screen "Dev_AI" 800x480, template "Settings"
   Softkey "Softkey_F3" at 0,0 size 0x0
      on KeyDown: function_dd21b452("AI_x_Result", 1)
   Softkey "Softkey_F7" at 0,0 size 0x0
      on KeyDown: SetBit("AI_x_CMD_Reset")
   Button "Button_2" at 165,265 size 112x32; TextOff 'DB 300'; Authorization "User administration"
      on Release: SetTag("AIx", 300); SetTag("AIx_Name", 'DB 300')
      Visibility <- "Support_DB_All_AIs"
      Appearance <- "AIx"
   Button "Button_8" at 165,305 size 112x32; TextOff 'DB 301'; Authorization "User administration"
      on Release: SetTag("AIx", 301); SetTag("AIx_Name", 'DB 301')
      Visibility <- "Support_DB_All_AIs"
      Appearance <- "AIx"
   Button "Button_17" at 165,345 size 112x32; TextOff 'DB 302'; Authorization "User administration"
      on Release: SetTag("AIx", 302); SetTag("AIx_Name", 'DB 302')
      Visibility <- "Support_DB_All_AIs"
      Appearance <- "AIx"
   Button "Button_18" at 165,385 size 112x32; TextOff 'DB 303'; Authorization "User administration"
      on Release: SetTag("AIx", 303); SetTag("AIx_Name", 'DB 303')
      Visibility <- "Support_DB_All_AIs"
      Appearance <- "AIx"
   Button "Button_3" at 443,265 size 112x32; TextOff 'DB 310'; Authorization "User administration"
      on Release: SetTag("AIx", 310); SetTag("AIx_Name", 'DB 310')
      Visibility <- "Support_DB_All_AIs"
      Appearance <- "AIx"
   Button "Button_4" at 443,305 size 112x32; TextOff 'DB 311'; Authorization "User administration"
      on Release: SetTag("AIx", 311); SetTag("AIx_Name", 'DB 311')
      Visibility <- "Support_DB_All_AIs"
      Appearance <- "AIx"
   Button "Button_6" at 443,345 size 112x32; TextOff 'DB 312'; Authorization "User administration"
      on Release: SetTag("AIx", 312); SetTag("AIx_Name", 'DB 312')
      Visibility <- "Support_DB_All_AIs"
      Appearance <- "AIx"
   Button "Button_10" at 443,385 size 112x32; TextOff 'DB 313'; Authorization "User administration"
      on Release: SetTag("AIx", 313); SetTag("AIx_Name", 'DB 313')
      Visibility <- "Support_DB_All_AIs"
      Appearance <- "AIx"
   Button "Button_11" at 443,425 size 112x32; TextOff 'DB 314'; Authorization "User administration"
      on Release: SetTag("AIx", 314); SetTag("AIx_Name", 'DB 314')
      Visibility <- "Support_DB_All_AIs"
      Appearance <- "AIx"
   Button "Button_1" at 583,344 size 112x32; TextOff 'DB 317'; Authorization "User administration"
      on Release: SetTag("AIx", 317); SetTag("AIx_Name", 'DB 317')
      Visibility <- "Support_DB_All_AIs"
      Appearance <- "AIx"
   Button "Button_5" at 583,384 size 112x32; TextOff 'DB 318'; Authorization "User administration"
      on Release: SetTag("AIx", 318); SetTag("AIx_Name", 'DB 318')
      Visibility <- "Support_DB_All_AIs"
      Appearance <- "AIx"
   Button "Button_9" at 583,264 size 112x32; TextOff 'DB 315'; Authorization "User administration"
      on Release: SetTag("AIx", 315); SetTag("AIx_Name", 'DB 315')
      Visibility <- "Support_DB_All_AIs"
      Appearance <- "AIx"
   Button "Button_14" at 583,304 size 112x32; TextOff 'DB 316'; Authorization "User administration"
      on Release: SetTag("AIx", 316); SetTag("AIx_Name", 'DB 316')
      Visibility <- "Support_DB_All_AIs"
      Appearance <- "AIx"
   Rectangle "Rectangle_3" at 165,7 size 530x150
      Appearance <- "AI_x_CMD_Start_A"
   Button "Button_7" at 171,43 size 80x22; TextOff 'Авто'; Authorization "User administration"; TextList "Hand"
      on Click: InvertBit("AI_x_CMD_Hand")
      Appearance <- "AI_x_CMD_Hand"
      ProcessValue <- "AI_x_CMD_Hand"
   TextField "Text field_1" at 484,12 size 107x18; Text 'Масштабирование'
      Visibility <- "AI_x_Use_RTD"
   TextField "Text field_20" at 495,24 size 18x18; Text 'от'
      Visibility <- "AI_x_Use_RTD"
   IOField "I/O field_5" at 476,42 size 65x20; Authorization "User administration"; FormatPattern 99999
      ProcessValue <- "AI_x_Converter_Min_In"
      Visibility <- "AI_x_Use_RTD"
   TextField "Text field_21" at 559,24 size 19x18; Text 'до'
      Visibility <- "AI_x_Use_RTD"
   IOField "I/O field_11" at 171,82 size 80x30; Authorization "User administration"; FormatPattern s9999.9
      ProcessValue <- "AI_x_Result"
      Appearance <- "AI_x_Status"
   TextField "Text field_22" at 177,64 size 68x18; Text 'Показания:'
   TextField "Text field_23" at 180,113 size 63x18; Text 'Вход ПЛК:'
   IOField "I/O field_17" at 171,133 size 80x20; FormatPattern s99999
      ProcessValue <- "AI_x_Signal"
   TextField "Text field_24" at 489,89 size 42x18; Text 'Обрыв'
      Visibility <- "AI_x_Alarm_NC"
   TextField "Text field_25" at 555,89 size 42x18; Text 'КЗ'
      Visibility <- "AI_x_Alarm_SC"
   IOField "I/O field_18" at 544,42 size 65x20; Authorization "User administration"; FormatPattern 99999
      ProcessValue <- "AI_x_Converter_Max_In"
      Visibility <- "AI_x_Use_RTD"
   IOField "I/O field_24" at 476,66 size 65x20; Authorization "User administration"; FormatPattern s9999.99
      ProcessValue <- "AI_x_Converter_Min_Out"
      Visibility <- "AI_x_Use_RTD"
   IOField "I/O field_25" at 544,66 size 65x20; Authorization "User administration"; FormatPattern s9999.99
      ProcessValue <- "AI_x_Converter_Max_Out"
      Visibility <- "AI_x_Use_RTD"
   IOField "I/O field_10" at 382,35 size 55x20; Authorization "User administration"; FormatPattern s9999.9
      Appearance <- "AI_x_Alarm_HH"
      ProcessValue <- "AI_x_SP_HH"
   TextField "Text field_10" at 354,36 size 28x18; Text 'HHS'
   TextField "Text field_12" at 354,60 size 20x18; Text 'HS'
   IOField "I/O field_12" at 382,58 size 55x20; Authorization "User administration"; FormatPattern s9999.9
      Appearance <- "AI_x_Alarm_H"
      ProcessValue <- "AI_x_SP_H"
   IOField "I/O field_26" at 440,35 size 26x20; Authorization "User administration"; FormatPattern 99.9
      Appearance <- "AI_x_Alarm_HH"
      ProcessValue <- "AI_x_Timers_HH_SP"
   IOField "I/O field_27" at 440,58 size 26x20; Authorization "User administration"; FormatPattern 99.9
      Appearance <- "AI_x_Alarm_H"
      ProcessValue <- "AI_x_Timers_H_SP"
   IOField "I/O field_28" at 382,82 size 55x20; Authorization "User administration"; FormatPattern s9999.9
      Appearance <- "AI_x_Alarm_L"
      ProcessValue <- "AI_x_SP_L"
   TextField "Text field_6" at 354,84 size 18x18; Text 'LS'
   TextField "Text field_28" at 354,108 size 24x18; Text 'LLS'
   IOField "I/O field_29" at 382,106 size 55x20; Authorization "User administration"; FormatPattern s9999.9
      Appearance <- "AI_x_Alarm_LL"
      ProcessValue <- "AI_x_SP_LL"
   IOField "I/O field_30" at 440,82 size 26x20; Authorization "User administration"; FormatPattern 99.9
      Appearance <- "AI_x_Alarm_L"
      ProcessValue <- "AI_x_Timers_L_SP"
   IOField "I/O field_31" at 440,106 size 26x20; Authorization "User administration"; FormatPattern 99.9
      Appearance <- "AI_x_Alarm_LL"
      ProcessValue <- "AI_x_Timers_LL_SP"
   IOField "I/O field_1" at 285,44 size 57x20; Authorization "Developer"; FormatPattern 999
      ProcessValue <- "AI_x_ADDR"
   TextField "Text field_2" at 262,45 size 21x18; Text 'IW'
   IOField "I/O field_8" at 171,12 size 171x26; FormatPattern ????????????????
      ProcessValue <- "AIx_Name"
   Button "Button_21" at 624,29 size 60x20; TextOff 'Text'; Authorization "User administration"; PictureList "Turn_ON"
      on Click: InvertBit("AI_x_Use_Filter")
      ProcessValue <- "AI_x_Use_Filter"
   TextField "Text field_3" at 616,11 size 75x18; Text 'Фильтрация'
   TextField "Text field_4" at 627,48 size 52x18; Text 'х0.1 сек'
   IOField "I/O field_2" at 624,67 size 60x20; Authorization "User administration"; FormatPattern 999
      ProcessValue <- "AI_x_Filter_SP"
   TextField "Text field_8" at 477,113 size 62x18; Text 'Поправка:'
   IOField "I/O field_3" at 549,111 size 60x20; Authorization "User administration"; FormatPattern s99.9
      ProcessValue <- "AI_x_Calibration"
   IOField "I/O field_4" at 568,133 size 44x20; Authorization "Developer"; FormatPattern 9999
      Visibility <- "AI_x_Use_RTD"
      ProcessValue <- "AI_x_RTD_c"
   TextField "Text field_11" at 267,64 size 81x18; Text 'Размерность:'
   TextField "Text field_13" at 275,113 size 67x18; Text 'Тип входа:'
   IOField "I/O field_6" at 264,133 size 42x20; Authorization "User administration"; FormatPattern 99.99
      ProcessValue <- "AI_x_VmA"
   Button "Button_19" at 266,82 size 80x30; TextOff 'Авто'; TextList "Input_Type"; Authorization "Developer"
      on Click: function_dd21b452("AI_x_Type", 1)
      ProcessValue <- "AI_x_Type"
   Button "Button_20" at 310,133 size 56x20; TextOff 'Авто'; Authorization "Developer"; TextList "VmA"
      on Click: function_dd21b452("AI_x_Input_Type", 1)
      ProcessValue <- "AI_x_Input_Type"
   TextField "Text field_14" at 348,12 size 123x18; Text 'Аварийные границы:'
   Button "Button_22" at 382,133 size 84x20; TextOff 'Сброс аварий'; Authorization "Operate"; TextList "VmA"
      on Click: SetBit("AI_x_CMD_Reset")
      ProcessValue <- "AI_x_CMD_Hand"
   Button "Button_24" at 170,130 size 82x24; TextOff 'Text'; Authorization "Developer"
      on Click: InvertBit("AI_x_CMD_Start_A")
   Button "Button_25" at 165,425 size 112x32; TextOff 'DB 304'; Authorization "User administration"
      on Release: SetTag("AIx", 304); SetTag("AIx_Name", 'DB 304')
      Visibility <- "Support_DB_All_AIs"
      Appearance <- "AIx"
   Button "Button_23" at 583,424 size 112x32; TextOff 'DB 319'; Authorization "User administration"
      on Release: SetTag("AIx", 319); SetTag("AIx_Name", 'DB 319')
      Visibility <- "Support_DB_All_AIs"
      Appearance <- "AIx"
   Button "Button_26" at 304,265 size 112x32; TextOff 'DB 305'; Authorization "User administration"
      on Release: SetTag("AIx", 305); SetTag("AIx_Name", 'DB 305')
      Visibility <- "Support_DB_All_AIs"
      Appearance <- "AIx"
   Button "Button_27" at 304,305 size 112x32; TextOff 'DB 306'; Authorization "User administration"
      on Release: SetTag("AIx", 306); SetTag("AIx_Name", 'DB 306')
      Visibility <- "Support_DB_All_AIs"
      Appearance <- "AIx"
   Button "Button_28" at 304,345 size 112x32; TextOff 'DB 307'; Authorization "User administration"
      on Release: SetTag("AIx", 307); SetTag("AIx_Name", 'DB 307')
      Visibility <- "Support_DB_All_AIs"
      Appearance <- "AIx"
   Button "Button_29" at 304,385 size 112x32; TextOff 'DB 308'; Authorization "User administration"
      on Release: SetTag("AIx", 308); SetTag("AIx_Name", 'DB 308')
      Visibility <- "Support_DB_All_AIs"
      Appearance <- "AIx"
   Button "Button_30" at 304,425 size 112x32; TextOff 'DB 309'; Authorization "User administration"
      on Release: SetTag("AIx", 309); SetTag("AIx_Name", 'DB 309')
      Visibility <- "Support_DB_All_AIs"
      Appearance <- "AIx"
   TextField "Text field_9" at 477,134 size 90x18; Text 'Коэффициент:'
      Visibility <- "AI_x_Use_RTD"
   Button "Button_12" at 624,108 size 60x20; TextOff 'Text'; PictureList "Turn_ON"; Authorization "User administration"
      on Click: InvertBit("AI_x_Use_Status")
      ProcessValue <- "AI_x_Use_Status"
   TextField "Text field_5" at 630,90 size 42x18; Text 'Статус'
   SymbolicIOField "Symbolic I/O field_1" at 113,464 size 75x16; TextOn '1'; TextOff '0'; TextList "Hand"
      ProcessValue <- "AI_x_CMD_Hand"
   TextField "Text field_7" at 211,464 size 75x16; Text 'Показания +1'
      Visibility <- "AI_x_CMD_Hand"
   TextField "Text field_15" at 311,464 size 75x16; Text 'Показания -1'
      Visibility <- "AI_x_CMD_Hand"
   TextField "Text field_16" at 610,464 size 75x16; Text 'Сброс аварий'
   Softkey "Softkey_F2" at 0,0 size 0x0
      on KeyDown: InvertBit("AI_x_CMD_Hand")
   Softkey "Softkey_F4" at 0,0 size 0x0
      on KeyDown: function_b9b71300("AI_x_Result", 1)

screen "Dev_DI_1" 800x480, template "Settings"
   TextField "Text field_4" at 134,11 size 130x26; Text 'Ав. Стоп'
   TextField "Text field_5" at 286,11 size 130x26; Text 'сигнал 2'
   TextField "Text field_29" at 438,11 size 130x26; Text 'сигнал 3'
   TextField "Text field_33" at 590,11 size 130x26; Text 'сигнал 4'
   TextField "Text field_17" at 134,283 size 130x26; Text 'сигнал 9'
   TextField "Text field_25" at 286,283 size 130x26; Text 'сигнал 10'
   TextField "Text field_9" at 134,147 size 130x26; Text 'сигнал 5'
   TextField "Text field_13" at 286,147 size 130x26; Text 'сигнал 6'
   TextField "Text field_21" at 438,147 size 130x26; Text 'сигнал 7'
   TextField "Text field_41" at 590,147 size 130x26; Text 'сигнал 8'
   TextField "Text field_37" at 590,283 size 130x26; Text 'сигнал 12'
   Button "Button_2" at 134,40 size 130x22; TextOff 'Авто'; Authorization "Operate"; TextList "Hand"
      on Click: InvertBit("DIx_Hand_x_1")
      Appearance <- "DIx_Hand_x_1"
      ProcessValue <- "DIx_Hand_x_1"
   Button "Button_3" at 204,65 size 60x20; TextOff 'Выкл'; Authorization "Operate"
      on Click: ResetBit("DIx_Start_M_x_1")
      Appearance <- "DIx_Start_M_x_1"
   Button "Button_13" at 134,65 size 60x20; TextOff 'Вкл'; Authorization "Operate"
      on Click: SetBit("DIx_Start_M_x_1")
      Appearance <- "DIx_Start_M_x_1"
   Button "Button_26" at 244,89 size 20x20; TextOff 'Text'; Authorization "User administration"; PictureList "ok_green"
      on Click: InvertBit("DIx_Inverse_x_1")
      ProcessValue <- "DIx_Inverse_x_1"
   TextField "Text field_1" at 133,85 size 91x23; Text 'Инверсия:'
   IOField "I/O field_1" at 176,109 size 30x24; Authorization "Developer"; FormatPattern 99
      ProcessValue <- "DIx_ADDR_Byte_x_1"
   IOField "I/O field_2" at 216,109 size 20x24; Authorization "Developer"; FormatPattern 9
      ProcessValue <- "DIx_ADDR_Bit_x_1"
   TextField "Text field_2" at 162,109 size 13x23; Text 'I'
   TextField "Text field_3" at 205,109 size 13x23; Text '.'
   Button "Button_1" at 286,40 size 130x22; TextOff 'Авто'; Authorization "Operate"; TextList "Hand"
      on Click: InvertBit("DIx_Hand_x_2")
      Appearance <- "DIx_Hand_x_2"
      ProcessValue <- "DIx_Hand_x_2"
   Button "Button_4" at 356,65 size 60x20; TextOff 'Выкл'; Authorization "Operate"
      on Click: ResetBit("DIx_Start_M_x_2")
      Appearance <- "DIx_Start_M_x_2"
   Button "Button_5" at 286,65 size 60x20; TextOff 'Вкл'; Authorization "Operate"
      on Click: SetBit("DIx_Start_M_x_2")
      Appearance <- "DIx_Start_M_x_2"
   Button "Button_6" at 396,89 size 20x20; TextOff 'Text'; Authorization "User administration"; PictureList "ok_green"
      on Click: InvertBit("DIx_Inverse_x_2")
      ProcessValue <- "DIx_Inverse_x_2"
   TextField "Text field_6" at 285,85 size 91x23; Text 'Инверсия:'
   IOField "I/O field_3" at 328,109 size 30x24; Authorization "Developer"; FormatPattern 99
      ProcessValue <- "DIx_ADDR_Byte_x_2"
   IOField "I/O field_4" at 368,109 size 20x24; Authorization "Developer"; FormatPattern 9
      ProcessValue <- "DIx_ADDR_Bit_x_2"
   TextField "Text field_7" at 314,109 size 13x23; Text 'I'
   TextField "Text field_8" at 357,109 size 13x23; Text '.'
   Button "Button_29" at 438,40 size 130x22; TextOff 'Авто'; Authorization "Operate"; TextList "Hand"
      on Click: InvertBit("DIx_Hand_x_3")
      Appearance <- "DIx_Hand_x_3"
      ProcessValue <- "DIx_Hand_x_3"
   Button "Button_30" at 508,65 size 60x20; TextOff 'Выкл'; Authorization "Operate"
      on Click: ResetBit("DIx_Start_M_x_3")
      Appearance <- "DIx_Start_M_x_3"
   Button "Button_31" at 438,65 size 60x20; TextOff 'Вкл'; Authorization "Operate"
      on Click: SetBit("DIx_Start_M_x_3")
      Appearance <- "DIx_Start_M_x_3"
   Button "Button_32" at 548,89 size 20x20; TextOff 'Text'; Authorization "User administration"; PictureList "ok_green"
      on Click: InvertBit("DIx_Inverse_x_3")
      ProcessValue <- "DIx_Inverse_x_3"
   TextField "Text field_30" at 437,85 size 91x23; Text 'Инверсия:'
   IOField "I/O field_15" at 480,109 size 30x24; Authorization "Developer"; FormatPattern 99
      ProcessValue <- "DIx_ADDR_Byte_x_3"
   IOField "I/O field_16" at 520,109 size 20x24; Authorization "Developer"; FormatPattern 9
      ProcessValue <- "DIx_ADDR_Bit_x_3"
   TextField "Text field_31" at 466,109 size 13x23; Text 'I'
   TextField "Text field_32" at 509,109 size 13x23; Text '.'
   Button "Button_7" at 590,40 size 130x22; TextOff 'Авто'; Authorization "Operate"; TextList "Hand"
      on Click: InvertBit("DIx_Hand_x_4")
      Appearance <- "DIx_Hand_x_4"
      ProcessValue <- "DIx_Hand_x_4"
   Button "Button_34" at 660,65 size 60x20; TextOff 'Выкл'; Authorization "Operate"
      on Click: ResetBit("DIx_Start_M_x_4")
      Appearance <- "DIx_Start_M_x_4"
   Button "Button_35" at 590,65 size 60x20; TextOff 'Вкл'; Authorization "Operate"
      on Click: SetBit("DIx_Start_M_x_4")
      Appearance <- "DIx_Start_M_x_4"
   Button "Button_36" at 700,89 size 20x20; TextOff 'Text'; Authorization "User administration"; PictureList "ok_green"
      on Click: InvertBit("DIx_Inverse_x_4")
      ProcessValue <- "DIx_Inverse_x_4"
   TextField "Text field_34" at 589,85 size 91x23; Text 'Инверсия:'
   IOField "I/O field_17" at 632,109 size 30x24; Authorization "Developer"; FormatPattern 99
      ProcessValue <- "DIx_ADDR_Byte_x_4"
   IOField "I/O field_18" at 672,109 size 20x24; Authorization "Developer"; FormatPattern 9
      ProcessValue <- "DIx_ADDR_Bit_x_4"
   TextField "Text field_35" at 618,109 size 13x23; Text 'I'
   TextField "Text field_36" at 661,109 size 13x23; Text '.'
   Button "Button_8" at 134,176 size 130x22; TextOff 'Авто'; Authorization "Operate"; TextList "Hand"
      on Click: InvertBit("DIx_Hand_x_5")
      Appearance <- "DIx_Hand_x_5"
      ProcessValue <- "DIx_Hand_x_5"
   Button "Button_9" at 204,201 size 60x20; TextOff 'Выкл'; Authorization "Operate"
      on Click: ResetBit("DIx_Start_M_x_5")
      Appearance <- "DIx_Start_M_x_5"
   Button "Button_10" at 134,201 size 60x20; TextOff 'Вкл'; Authorization "Operate"
      on Click: SetBit("DIx_Start_M_x_5")
      Appearance <- "DIx_Start_M_x_5"
   Button "Button_11" at 244,225 size 20x20; TextOff 'Text'; Authorization "User administration"; PictureList "ok_green"
      on Click: InvertBit("DIx_Inverse_x_5")
      ProcessValue <- "DIx_Inverse_x_5"
   TextField "Text field_10" at 133,221 size 91x23; Text 'Инверсия:'
   IOField "I/O field_5" at 176,245 size 30x24; Authorization "Developer"; FormatPattern 99
      ProcessValue <- "DIx_ADDR_Byte_x_5"
   IOField "I/O field_6" at 216,245 size 20x24; Authorization "Developer"; FormatPattern 9
      ProcessValue <- "DIx_ADDR_Bit_x_5"
   TextField "Text field_11" at 162,245 size 13x23; Text 'I'
   TextField "Text field_12" at 205,245 size 13x23; Text '.'
   Button "Button_12" at 286,176 size 130x22; TextOff 'Авто'; Authorization "Operate"; TextList "Hand"
      on Click: InvertBit("DIx_Hand_x_6")
      Appearance <- "DIx_Hand_x_6"
      ProcessValue <- "DIx_Hand_x_6"
   Button "Button_14" at 356,201 size 60x20; TextOff 'Выкл'; Authorization "Operate"
      on Click: ResetBit("DIx_Start_M_x_6")
      Appearance <- "DIx_Start_M_x_6"
   Button "Button_15" at 286,201 size 60x20; TextOff 'Вкл'; Authorization "Operate"
      on Click: SetBit("DIx_Start_M_x_6")
      Appearance <- "DIx_Start_M_x_6"
   Button "Button_16" at 396,225 size 20x20; TextOff 'Text'; Authorization "User administration"; PictureList "ok_green"
      on Click: InvertBit("DIx_Inverse_x_6")
      ProcessValue <- "DIx_Inverse_x_6"
   TextField "Text field_14" at 285,221 size 91x23; Text 'Инверсия:'
   IOField "I/O field_7" at 328,245 size 30x24; Authorization "Developer"; FormatPattern 99
      ProcessValue <- "DIx_ADDR_Byte_x_6"
   IOField "I/O field_8" at 368,245 size 20x24; Authorization "Developer"; FormatPattern 9
      ProcessValue <- "DIx_ADDR_Bit_x_6"
   TextField "Text field_15" at 314,245 size 13x23; Text 'I'
   TextField "Text field_16" at 357,245 size 13x23; Text '.'
   Button "Button_20" at 438,176 size 130x22; TextOff 'Авто'; Authorization "Operate"; TextList "Hand"
      on Click: InvertBit("DIx_Hand_x_7")
      Appearance <- "DIx_Hand_x_7"
      ProcessValue <- "DIx_Hand_x_7"
   Button "Button_21" at 508,201 size 60x20; TextOff 'Выкл'; Authorization "Operate"
      on Click: ResetBit("DIx_Start_M_x_7")
      Appearance <- "DIx_Start_M_x_7"
   Button "Button_22" at 438,201 size 60x20; TextOff 'Вкл'; Authorization "Operate"
      on Click: SetBit("DIx_Start_M_x_7")
      Appearance <- "DIx_Start_M_x_7"
   Button "Button_23" at 548,225 size 20x20; TextOff 'Text'; Authorization "User administration"; PictureList "ok_green"
      on Click: InvertBit("DIx_Inverse_x_7")
      ProcessValue <- "DIx_Inverse_x_7"
   TextField "Text field_22" at 437,221 size 91x23; Text 'Инверсия:'
   IOField "I/O field_11" at 480,245 size 30x24; Authorization "Developer"; FormatPattern 99
      ProcessValue <- "DIx_ADDR_Byte_x_7"
   IOField "I/O field_12" at 520,245 size 20x24; Authorization "Developer"; FormatPattern 9
      ProcessValue <- "DIx_ADDR_Bit_x_7"
   TextField "Text field_23" at 466,245 size 13x23; Text 'I'
   TextField "Text field_24" at 509,245 size 13x23; Text '.'
   Button "Button_41" at 590,176 size 130x22; TextOff 'Авто'; Authorization "Operate"; TextList "Hand"
      on Click: InvertBit("DIx_Hand_x_8")
      Appearance <- "DIx_Hand_x_8"
      ProcessValue <- "DIx_Hand_x_8"
   Button "Button_42" at 660,201 size 60x20; TextOff 'Выкл'; Authorization "Operate"
      on Click: ResetBit("DIx_Start_M_x_8")
      Appearance <- "DIx_Start_M_x_8"
   Button "Button_43" at 590,201 size 60x20; TextOff 'Вкл'; Authorization "Operate"
      on Click: SetBit("DIx_Start_M_x_8")
      Appearance <- "DIx_Start_M_x_8"
   Button "Button_44" at 700,225 size 20x20; TextOff 'Text'; Authorization "User administration"; PictureList "ok_green"
      on Click: InvertBit("DIx_Inverse_x_8")
      ProcessValue <- "DIx_Inverse_x_8"
   TextField "Text field_42" at 589,221 size 91x23; Text 'Инверсия:'
   IOField "I/O field_21" at 632,245 size 30x24; Authorization "Developer"; FormatPattern 99
      ProcessValue <- "DIx_ADDR_Byte_x_8"
   IOField "I/O field_22" at 672,245 size 20x24; Authorization "Developer"; FormatPattern 9
      ProcessValue <- "DIx_ADDR_Bit_x_8"
   TextField "Text field_43" at 618,245 size 13x23; Text 'I'
   TextField "Text field_44" at 661,245 size 13x23; Text '.'
   Button "Button_24" at 134,312 size 130x22; TextOff 'Авто'; Authorization "Operate"; TextList "Hand"
      on Click: InvertBit("DIx_Hand_x_9")
      Appearance <- "DIx_Hand_x_9"
      ProcessValue <- "DIx_Hand_x_9"
   Button "Button_25" at 204,337 size 60x20; TextOff 'Выкл'; Authorization "Operate"
      on Click: ResetBit("DIx_Start_M_x_9")
      Appearance <- "DIx_Start_M_x_9"
   Button "Button_27" at 134,337 size 60x20; TextOff 'Вкл'; Authorization "Operate"
      on Click: SetBit("DIx_Start_M_x_9")
      Appearance <- "DIx_Start_M_x_9"
   Button "Button_28" at 244,361 size 20x20; TextOff 'Text'; Authorization "User administration"; PictureList "ok_green"
      on Click: InvertBit("DIx_Inverse_x_9")
      ProcessValue <- "DIx_Inverse_x_9"
   TextField "Text field_18" at 133,357 size 91x23; Text 'Инверсия:'
   IOField "I/O field_9" at 176,381 size 30x24; Authorization "Developer"; FormatPattern 99
      ProcessValue <- "DIx_ADDR_Byte_x_9"
   IOField "I/O field_10" at 216,381 size 20x24; Authorization "Developer"; FormatPattern 9
      ProcessValue <- "DIx_ADDR_Bit_x_9"
   TextField "Text field_19" at 162,381 size 13x23; Text 'I'
   TextField "Text field_20" at 205,381 size 13x23; Text '.'
   Button "Button_37" at 286,312 size 130x22; TextOff 'Авто'; Authorization "Operate"; TextList "Hand"
      on Click: InvertBit("DIx_Hand_x_10")
      Appearance <- "DIx_Hand_x_10"
      ProcessValue <- "DIx_Hand_x_10"
   Button "Button_38" at 356,337 size 60x20; TextOff 'Выкл'; Authorization "Operate"
      on Click: ResetBit("DIx_Start_M_x_10")
      Appearance <- "DIx_Start_M_x_10"
   Button "Button_39" at 286,337 size 60x20; TextOff 'Вкл'; Authorization "Operate"
      on Click: SetBit("DIx_Start_M_x_10")
      Appearance <- "DIx_Start_M_x_10"
   Button "Button_40" at 396,361 size 20x20; TextOff 'Text'; Authorization "User administration"; PictureList "ok_green"
      on Click: InvertBit("DIx_Inverse_x_10")
      ProcessValue <- "DIx_Inverse_x_10"
   TextField "Text field_26" at 285,357 size 91x23; Text 'Инверсия:'
   IOField "I/O field_13" at 328,381 size 30x24; Authorization "Developer"; FormatPattern 99
      ProcessValue <- "DIx_ADDR_Byte_x_10"
   IOField "I/O field_14" at 368,381 size 20x24; Authorization "Developer"; FormatPattern 9
      ProcessValue <- "DIx_ADDR_Bit_x_10"
   TextField "Text field_27" at 314,381 size 13x23; Text 'I'
   TextField "Text field_28" at 357,381 size 13x23; Text '.'
   Button "Button_48" at 590,312 size 130x22; TextOff 'Авто'; Authorization "Operate"; TextList "Hand"
      on Click: InvertBit("DIx_Hand_x_12")
      Appearance <- "DIx_Hand_x_12"
      ProcessValue <- "DIx_Hand_x_12"
   Button "Button_49" at 660,337 size 60x20; TextOff 'Выкл'; Authorization "Operate"
      on Click: ResetBit("DIx_Start_M_x_12")
      Appearance <- "DIx_Start_M_x_12"
   Button "Button_50" at 590,337 size 60x20; TextOff 'Вкл'; Authorization "Operate"
      on Click: SetBit("DIx_Start_M_x_12")
      Appearance <- "DIx_Start_M_x_12"
   Button "Button_51" at 700,361 size 20x20; TextOff 'Text'; Authorization "User administration"; PictureList "ok_green"
      on Click: InvertBit("DIx_Inverse_x_12")
      ProcessValue <- "DIx_Inverse_x_12"
   TextField "Text field_45" at 589,357 size 91x23; Text 'Инверсия:'
   IOField "I/O field_23" at 632,381 size 30x24; Authorization "Developer"; FormatPattern 99
      ProcessValue <- "DIx_ADDR_Byte_x_12"
   IOField "I/O field_24" at 672,381 size 20x24; Authorization "Developer"; FormatPattern 9
      ProcessValue <- "DIx_ADDR_Bit_x_12"
   TextField "Text field_46" at 618,381 size 13x23; Text 'I'
   TextField "Text field_47" at 661,381 size 13x23; Text '.'
   TextField "Text field_38" at 438,283 size 130x26; Text 'сигнал 11'
   Button "Button_17" at 438,312 size 130x22; TextOff 'Авто'; Authorization "Operate"; TextList "Hand"
      on Click: InvertBit("DIx_Hand_x_11")
      Appearance <- "DIx_Hand_x_11"
      ProcessValue <- "DIx_Hand_x_11"
   Button "Button_18" at 508,337 size 60x20; TextOff 'Выкл'; Authorization "Operate"
      on Click: ResetBit("DIx_Start_M_x_11")
      Appearance <- "DIx_Start_M_x_11"
   Button "Button_19" at 438,337 size 60x20; TextOff 'Вкл'; Authorization "Operate"
      on Click: SetBit("DIx_Start_M_x_11")
      Appearance <- "DIx_Start_M_x_11"
   Button "Button_52" at 548,361 size 20x20; TextOff 'Text'; Authorization "User administration"; PictureList "ok_green"
      on Click: InvertBit("DIx_Inverse_x_11")
      ProcessValue <- "DIx_Inverse_x_11"
   TextField "Text field_39" at 437,357 size 91x23; Text 'Инверсия:'
   IOField "I/O field_19" at 480,381 size 30x24; Authorization "Developer"; FormatPattern 99
      ProcessValue <- "DIx_ADDR_Byte_x_11"
   IOField "I/O field_20" at 520,381 size 20x24; Authorization "Developer"; FormatPattern 9
      ProcessValue <- "DIx_ADDR_Bit_x_11"
   TextField "Text field_40" at 466,381 size 13x23; Text 'I'
   TextField "Text field_48" at 509,381 size 13x23; Text '.'
   Button "Button_33" at 128,440 size 75x30; TextOff 'Стр.1'; Authorization "Operate"
      on Click: SetTag("DIx", 200); ActivateScreen("Dev_DI_1", 0)
      Visibility <- "Support_DB_All_DIs"
      Appearance <- "DIx"
   Button "Button_45" at 233,440 size 75x30; TextOff 'Стр.2'; Authorization "Operate"
      on Click: SetTag("DIx", 201); ActivateScreen("Dev_DI_2", 0)
      Visibility <- "Support_DB_All_DIs"
      Appearance <- "DIx"
   Button "Button_46" at 338,440 size 75x30; TextOff 'Стр.3'; Authorization "Operate"
      on Click: SetTag("DIx", 202); ActivateScreen("Dev_DI_3", 0)
      Visibility <- "Support_DB_All_DIs"
      Appearance <- "DIx"
   Button "Button_47" at 444,440 size 75x30; TextOff 'Стр.4'; Authorization "Operate"
      on Click: SetTag("DIx", 203); ActivateScreen("Dev_DI_4", 0)
      Visibility <- "Support_DB_All_DIs"
      Appearance <- "DIx"
   Button "Button_53" at 549,440 size 75x30; TextOff 'Стр.5'; Authorization "Operate"
      on Click: SetTag("DIx", 204); ActivateScreen("Dev_DI_5", 0)
      Visibility <- "Support_DB_All_DIs"
      Appearance <- "DIx"
   Button "Button_54" at 655,440 size 75x30; TextOff 'Стр.6'; Authorization "Operate"
      on Click: SetTag("DIx", 205); ActivateScreen("Dev_DI_6", 0)
      Visibility <- "Support_DB_All_DIs"
      Appearance <- "DIx"

screen "Dev_DO_1" 800x480, template "Settings"
   TextField "Text field_4" at 134,11 size 130x26; Text 'выход 1'
   TextField "Text field_5" at 286,11 size 130x26; Text 'выход 2'
   TextField "Text field_29" at 438,11 size 130x26; Text 'выход 3'
   TextField "Text field_33" at 590,11 size 130x26; Text 'выход 4'
   TextField "Text field_17" at 134,283 size 130x26; Text 'выход 9'
   TextField "Text field_25" at 286,283 size 130x26; Text 'выход 10'
   TextField "Text field_9" at 134,147 size 130x26; Text 'выход 5'
   TextField "Text field_13" at 286,147 size 130x26; Text 'выход 6'
   TextField "Text field_21" at 438,147 size 130x26; Text 'выход 7'
   TextField "Text field_41" at 590,147 size 130x26; Text 'выход 8'
   TextField "Text field_37" at 590,283 size 130x26; Text 'выход 12'
   Button "Button_2" at 134,40 size 130x22; TextOff 'Авто'; Authorization "Operate"; TextList "Hand"
      on Click: InvertBit("DOx_Hand_x_1")
      Appearance <- "DOx_Hand_x_1"
      ProcessValue <- "DOx_Hand_x_1"
   Button "Button_13" at 134,65 size 60x20; TextOff 'Вкл'; Authorization "Operate"
      on Click: SetBit("DOx_Start_M_x_1")
      Appearance <- "DOx_Start_M_x_1"
   Button "Button_26" at 244,89 size 20x20; TextOff 'Text'; PictureList "ok_green"; Authorization "User administration"
      on Click: InvertBit("DOx_Inverse_x_1")
      ProcessValue <- "DOx_Inverse_x_1"
   TextField "Text field_1" at 133,85 size 91x23; Text 'Инверсия:'
   IOField "I/O field_1" at 176,109 size 30x24; Authorization "Developer"; FormatPattern 99
      ProcessValue <- "DOx_ADDR_Byte_x_1"
   IOField "I/O field_2" at 216,109 size 20x24; Authorization "Developer"; FormatPattern 9
      ProcessValue <- "DOx_ADDR_Bit_x_1"
   TextField "Text field_2" at 158,109 size 20x23; Text 'Q'
   TextField "Text field_3" at 205,109 size 13x23; Text '.'
   Button "Button_1" at 286,40 size 130x22; TextOff 'Авто'; Authorization "Operate"; TextList "Hand"
      on Click: InvertBit("DOx_Hand_x_2")
      Appearance <- "DOx_Hand_x_2"
      ProcessValue <- "DOx_Hand_x_2"
   Button "Button_5" at 286,65 size 60x20; TextOff 'Вкл'; Authorization "Operate"
      on Click: SetBit("DOx_Start_M_x_2")
      Appearance <- "DOx_Start_M_x_2"
   Button "Button_6" at 396,89 size 20x20; TextOff 'Text'; Authorization "User administration"; PictureList "ok_green"
      on Click: InvertBit("DOx_Inverse_x_2")
      ProcessValue <- "DOx_Inverse_x_2"
   TextField "Text field_6" at 285,85 size 91x23; Text 'Инверсия:'
   IOField "I/O field_3" at 328,109 size 30x24; Authorization "Developer"; FormatPattern 99
      ProcessValue <- "DOx_ADDR_Byte_x_2"
   IOField "I/O field_4" at 368,109 size 20x24; Authorization "Developer"; FormatPattern 9
      ProcessValue <- "DOx_ADDR_Bit_x_2"
   TextField "Text field_7" at 310,109 size 20x23; Text 'Q'
   TextField "Text field_8" at 357,109 size 13x23; Text '.'
   Button "Button_29" at 438,40 size 130x22; TextOff 'Авто'; Authorization "Operate"; TextList "Hand"
      on Click: InvertBit("DOx_Hand_x_3")
      Appearance <- "DOx_Hand_x_3"
      ProcessValue <- "DOx_Hand_x_3"
   Button "Button_31" at 438,65 size 60x20; TextOff 'Вкл'; Authorization "Operate"
      on Click: SetBit("DOx_Start_M_x_3")
      Appearance <- "DOx_Start_M_x_3"
   Button "Button_32" at 548,89 size 20x20; TextOff 'Text'; Authorization "User administration"; PictureList "ok_green"
      on Click: InvertBit("DOx_Inverse_x_3")
      ProcessValue <- "DOx_Inverse_x_3"
   TextField "Text field_30" at 437,85 size 91x23; Text 'Инверсия:'
   IOField "I/O field_15" at 480,109 size 30x24; Authorization "Developer"; FormatPattern 99
      ProcessValue <- "DOx_ADDR_Byte_x_3"
   IOField "I/O field_16" at 520,109 size 20x24; Authorization "Developer"; FormatPattern 9
      ProcessValue <- "DOx_ADDR_Bit_x_3"
   TextField "Text field_31" at 462,109 size 20x23; Text 'Q'
   TextField "Text field_32" at 509,109 size 13x23; Text '.'
   Button "Button_33" at 590,40 size 130x22; TextOff 'Авто'; Authorization "Operate"; TextList "Hand"
      on Click: InvertBit("DOx_Hand_x_4")
      Appearance <- "DOx_Hand_x_4"
      ProcessValue <- "DOx_Hand_x_4"
   Button "Button_35" at 590,65 size 60x20; TextOff 'Вкл'; Authorization "Operate"
      on Click: SetBit("DOx_Start_M_x_4")
      Appearance <- "DOx_Start_M_x_4"
   Button "Button_36" at 700,89 size 20x20; TextOff 'Text'; Authorization "User administration"; PictureList "ok_green"
      on Click: InvertBit("DOx_Inverse_x_4")
      ProcessValue <- "DOx_Inverse_x_4"
   TextField "Text field_34" at 589,85 size 91x23; Text 'Инверсия:'
   IOField "I/O field_17" at 632,109 size 30x24; Authorization "Developer"; FormatPattern 99
      ProcessValue <- "DOx_ADDR_Byte_x_4"
   IOField "I/O field_18" at 672,109 size 20x24; Authorization "Developer"; FormatPattern 9
      ProcessValue <- "DOx_ADDR_Bit_x_4"
   TextField "Text field_35" at 614,109 size 20x23; Text 'Q'
   TextField "Text field_36" at 661,109 size 13x23; Text '.'
   Button "Button_7" at 134,176 size 130x22; TextOff 'Авто'; Authorization "Operate"; TextList "Hand"
      on Click: InvertBit("DOx_Hand_x_5")
      Appearance <- "DOx_Hand_x_5"
      ProcessValue <- "DOx_Hand_x_5"
   Button "Button_9" at 134,201 size 60x20; TextOff 'Вкл'; Authorization "Operate"
      on Click: SetBit("DOx_Start_M_x_5")
      Appearance <- "DOx_Start_M_x_5"
   Button "Button_10" at 244,225 size 20x20; TextOff 'Text'; Authorization "User administration"; PictureList "ok_green"
      on Click: InvertBit("DOx_Inverse_x_5")
      ProcessValue <- "DOx_Inverse_x_5"
   TextField "Text field_10" at 133,221 size 91x23; Text 'Инверсия:'
   IOField "I/O field_5" at 176,245 size 30x24; Authorization "Developer"; FormatPattern 99
      ProcessValue <- "DOx_ADDR_Byte_x_5"
   IOField "I/O field_6" at 216,245 size 20x24; Authorization "Developer"; FormatPattern 9
      ProcessValue <- "DOx_ADDR_Bit_x_5"
   TextField "Text field_11" at 158,245 size 20x23; Text 'Q'
   TextField "Text field_12" at 205,245 size 13x23; Text '.'
   Button "Button_11" at 286,176 size 130x22; TextOff 'Авто'; Authorization "Operate"; TextList "Hand"
      on Click: InvertBit("DOx_Hand_x_6")
      Appearance <- "DOx_Hand_x_6"
      ProcessValue <- "DOx_Hand_x_6"
   Button "Button_14" at 286,201 size 60x20; TextOff 'Вкл'; Authorization "Operate"
      on Click: SetBit("DOx_Start_M_x_6")
      Appearance <- "DOx_Start_M_x_6"
   Button "Button_15" at 396,225 size 20x20; TextOff 'Text'; PictureList "ok_green"; Authorization "User administration"
      on Click: InvertBit("DOx_Inverse_x_6")
      ProcessValue <- "DOx_Inverse_x_6"
   TextField "Text field_14" at 285,221 size 91x23; Text 'Инверсия:'
   IOField "I/O field_7" at 328,245 size 30x24; Authorization "Developer"; FormatPattern 99
      ProcessValue <- "DOx_ADDR_Byte_x_6"
   IOField "I/O field_8" at 368,245 size 20x24; Authorization "Developer"; FormatPattern 9
      ProcessValue <- "DOx_ADDR_Bit_x_6"
   TextField "Text field_15" at 310,245 size 20x23; Text 'Q'
   TextField "Text field_16" at 357,245 size 13x23; Text '.'
   Button "Button_20" at 438,176 size 130x22; TextOff 'Авто'; Authorization "Operate"; TextList "Hand"
      on Click: InvertBit("DOx_Hand_x_7")
      Appearance <- "DOx_Hand_x_7"
      ProcessValue <- "DOx_Hand_x_7"
   Button "Button_22" at 438,201 size 60x20; TextOff 'Вкл'; Authorization "Operate"
      on Click: SetBit("DOx_Start_M_x_7")
      Appearance <- "DOx_Start_M_x_7"
   Button "Button_23" at 548,225 size 20x20; TextOff 'Text'; PictureList "ok_green"; Authorization "User administration"
      on Click: InvertBit("DOx_Inverse_x_7")
      ProcessValue <- "DOx_Inverse_x_7"
   TextField "Text field_22" at 437,221 size 91x23; Text 'Инверсия:'
   IOField "I/O field_11" at 480,245 size 30x24; Authorization "Developer"; FormatPattern 99
      ProcessValue <- "DOx_ADDR_Byte_x_7"
   IOField "I/O field_12" at 520,245 size 20x24; Authorization "Developer"; FormatPattern 9
      ProcessValue <- "DOx_ADDR_Bit_x_7"
   TextField "Text field_23" at 462,245 size 20x23; Text 'Q'
   TextField "Text field_24" at 509,245 size 13x23; Text '.'
   Button "Button_41" at 590,176 size 130x22; TextOff 'Авто'; Authorization "Operate"; TextList "Hand"
      on Click: InvertBit("DOx_Hand_x_8")
      Appearance <- "DOx_Hand_x_8"
      ProcessValue <- "DOx_Hand_x_8"
   Button "Button_43" at 590,201 size 60x20; TextOff 'Вкл'; Authorization "Operate"
      on Click: SetBit("DOx_Start_M_x_8")
      Appearance <- "DOx_Start_M_x_8"
   Button "Button_44" at 700,225 size 20x20; TextOff 'Text'; PictureList "ok_green"; Authorization "User administration"
      on Click: InvertBit("DOx_Inverse_x_8")
      ProcessValue <- "DOx_Inverse_x_8"
   TextField "Text field_42" at 589,221 size 91x23; Text 'Инверсия:'
   IOField "I/O field_21" at 632,245 size 30x24; Authorization "Developer"; FormatPattern 99
      ProcessValue <- "DOx_ADDR_Byte_x_8"
   IOField "I/O field_22" at 672,245 size 20x24; Authorization "Developer"; FormatPattern 9
      ProcessValue <- "DOx_ADDR_Bit_x_8"
   TextField "Text field_43" at 614,245 size 20x23; Text 'Q'
   TextField "Text field_44" at 661,245 size 13x23; Text '.'
   Button "Button_24" at 134,312 size 130x22; TextOff 'Авто'; Authorization "Operate"; TextList "Hand"
      on Click: InvertBit("DOx_Hand_x_9")
      Appearance <- "DOx_Hand_x_9"
      ProcessValue <- "DOx_Hand_x_9"
   Button "Button_27" at 134,337 size 60x20; TextOff 'Вкл'; Authorization "Operate"
      on Click: SetBit("DOx_Start_M_x_9")
      Appearance <- "DOx_Start_M_x_9"
   Button "Button_28" at 244,361 size 20x20; TextOff 'Text'; Authorization "User administration"; PictureList "ok_green"
      on Click: InvertBit("DOx_Inverse_x_9")
      ProcessValue <- "DOx_Inverse_x_9"
   TextField "Text field_18" at 133,357 size 91x23; Text 'Инверсия:'
   IOField "I/O field_9" at 176,381 size 30x24; Authorization "Developer"; FormatPattern 99
      ProcessValue <- "DOx_ADDR_Byte_x_9"
   IOField "I/O field_10" at 216,381 size 20x24; Authorization "Developer"; FormatPattern 9
      ProcessValue <- "DOx_ADDR_Bit_x_9"
   TextField "Text field_19" at 158,381 size 20x23; Text 'Q'
   TextField "Text field_20" at 205,381 size 13x23; Text '.'
   Button "Button_37" at 286,312 size 130x22; TextOff 'Авто'; Authorization "Operate"; TextList "Hand"
      on Click: InvertBit("DOx_Hand_x_10")
      Appearance <- "DOx_Hand_x_10"
      ProcessValue <- "DOx_Hand_x_10"
   Button "Button_39" at 286,337 size 60x20; TextOff 'Вкл'; Authorization "Operate"
      on Click: SetBit("DOx_Start_M_x_10")
      Appearance <- "DOx_Start_M_x_10"
   Button "Button_40" at 396,361 size 20x20; TextOff 'Text'; PictureList "ok_green"; Authorization "User administration"
      on Click: InvertBit("DOx_Inverse_x_10")
      ProcessValue <- "DOx_Inverse_x_10"
   TextField "Text field_26" at 285,357 size 91x23; Text 'Инверсия:'
   IOField "I/O field_13" at 328,381 size 30x24; Authorization "Developer"; FormatPattern 99
      ProcessValue <- "DOx_ADDR_Byte_x_10"
   IOField "I/O field_14" at 368,381 size 20x24; Authorization "Developer"; FormatPattern 9
      ProcessValue <- "DOx_ADDR_Bit_x_10"
   TextField "Text field_27" at 310,381 size 20x23; Text 'Q'
   TextField "Text field_28" at 357,381 size 13x23; Text '.'
   Button "Button_48" at 590,312 size 130x22; TextOff 'Авто'; Authorization "Operate"; TextList "Hand"
      on Click: InvertBit("DOx_Hand_x_12")
      Appearance <- "DOx_Hand_x_12"
      ProcessValue <- "DOx_Hand_x_12"
   Button "Button_50" at 590,337 size 60x20; TextOff 'Вкл'; Authorization "Operate"
      on Click: SetBit("DOx_Start_M_x_12")
      Appearance <- "DOx_Start_M_x_12"
   Button "Button_51" at 700,361 size 20x20; TextOff 'Text'; PictureList "ok_green"; Authorization "User administration"
      on Click: InvertBit("DOx_Inverse_x_12")
      ProcessValue <- "DOx_Inverse_x_12"
   TextField "Text field_45" at 589,357 size 91x23; Text 'Инверсия:'
   IOField "I/O field_23" at 632,381 size 30x24; Authorization "Developer"; FormatPattern 99
      ProcessValue <- "DOx_ADDR_Byte_x_12"
   IOField "I/O field_24" at 672,381 size 20x24; Authorization "Developer"; FormatPattern 9
      ProcessValue <- "DOx_ADDR_Bit_x_12"
   TextField "Text field_46" at 614,381 size 20x23; Text 'Q'
   TextField "Text field_47" at 661,381 size 13x23; Text '.'
   TextField "Text field_38" at 438,283 size 130x26; Text 'выход 11'
   Button "Button_45" at 438,312 size 130x22; TextOff 'Авто'; Authorization "Operate"; TextList "Hand"
      on Click: InvertBit("DOx_Hand_x_11")
      Appearance <- "DOx_Hand_x_11"
      ProcessValue <- "DOx_Hand_x_11"
   Button "Button_47" at 438,337 size 60x20; TextOff 'Вкл'; Authorization "Operate"
      on Click: SetBit("DOx_Start_M_x_11")
      Appearance <- "DOx_Start_M_x_11"
   Button "Button_52" at 548,361 size 20x20; TextOff 'Text'; Authorization "User administration"; PictureList "ok_green"
      on Click: InvertBit("DOx_Inverse_x_11")
      ProcessValue <- "DOx_Inverse_x_11"
   TextField "Text field_39" at 437,357 size 91x23; Text 'Инверсия:'
   IOField "I/O field_19" at 480,381 size 30x24; Authorization "Developer"; FormatPattern 99
      ProcessValue <- "DOx_ADDR_Byte_x_11"
   IOField "I/O field_20" at 520,381 size 20x24; Authorization "Developer"; FormatPattern 9
      ProcessValue <- "DOx_ADDR_Bit_x_11"
   TextField "Text field_40" at 462,381 size 20x23; Text 'Q'
   TextField "Text field_48" at 509,381 size 13x23; Text '.'
   Button "Button_16" at 128,440 size 75x30; TextOff 'Стр.1'; Authorization "Operate"
      on Click: SetTag("DOx", 210); ActivateScreen("Dev_DI_1", 0)
      Visibility <- "Support_DB_All_DOs"
      Appearance <- "DOx"
   Button "Button_17" at 233,440 size 75x30; TextOff 'Стр.2'; Authorization "Operate"
      on Click: SetTag("DOx", 211); ActivateScreen("Dev_DI_2", 0)
      Visibility <- "Support_DB_All_DOs"
      Appearance <- "DOx"
   Button "Button_18" at 338,440 size 75x30; TextOff 'Стр.3'; Authorization "Operate"
      on Click: SetTag("DOx", 212); ActivateScreen("Dev_DI_3", 0)
      Visibility <- "Support_DB_All_DOs"
      Appearance <- "DOx"
   Button "Button_19" at 444,440 size 75x30; TextOff 'Стр.4'; Authorization "Operate"
      on Click: SetTag("DOx", 213); ActivateScreen("Dev_DI_4", 0)
      Visibility <- "Support_DB_All_DOs"
      Appearance <- "DOx"
   Button "Button_53" at 549,440 size 75x30; TextOff 'Стр.5'; Authorization "Operate"
      on Click: SetTag("DOx", 214); ActivateScreen("Dev_DI_5", 0)
      Visibility <- "Support_DB_All_DOs"
      Appearance <- "DOx"
   Button "Button_54" at 655,440 size 75x30; TextOff 'Стр.6'; Authorization "Operate"
      on Click: SetTag("DOx", 215); ActivateScreen("Dev_DI_6", 0)
      Visibility <- "Support_DB_All_DOs"
      Appearance <- "DOx"
   Button "Button_3" at 204,65 size 60x20; TextOff 'Выкл'; Authorization "Operate"
      on Click: ResetBit("DOx_Start_M_x_1")
      Appearance <- "DOx_Start_M_x_1"
   Button "Button_4" at 356,65 size 60x20; TextOff 'Выкл'; Authorization "Operate"
      on Click: ResetBit("DOx_Start_M_x_2")
      Appearance <- "DOx_Start_M_x_2"
   Button "Button_30" at 508,65 size 60x20; TextOff 'Выкл'; Authorization "Operate"
      on Click: ResetBit("DOx_Start_M_x_3")
      Appearance <- "DOx_Start_M_x_3"
   Button "Button_34" at 660,65 size 60x20; TextOff 'Выкл'; Authorization "Operate"
      on Click: ResetBit("DOx_Start_M_x_4")
      Appearance <- "DOx_Start_M_x_4"
   Button "Button_8" at 204,201 size 60x20; TextOff 'Выкл'; Authorization "Operate"
      on Click: ResetBit("DOx_Start_M_x_5")
      Appearance <- "DOx_Start_M_x_5"
   Button "Button_12" at 356,201 size 60x20; TextOff 'Выкл'; Authorization "Operate"
      on Click: ResetBit("DOx_Start_M_x_6")
      Appearance <- "DOx_Start_M_x_6"
   Button "Button_21" at 508,201 size 60x20; TextOff 'Выкл'; Authorization "Operate"
      on Click: ResetBit("DOx_Start_M_x_7")
      Appearance <- "DOx_Start_M_x_7"
   Button "Button_42" at 660,201 size 60x20; TextOff 'Выкл'; Authorization "Operate"
      on Click: ResetBit("DOx_Start_M_x_8")
      Appearance <- "DOx_Start_M_x_8"
   Button "Button_25" at 204,337 size 60x20; TextOff 'Выкл'; Authorization "Operate"
      on Click: ResetBit("DOx_Start_M_x_9")
      Appearance <- "DOx_Start_M_x_9"
   Button "Button_38" at 356,337 size 60x20; TextOff 'Выкл'; Authorization "Operate"
      on Click: ResetBit("DOx_Start_M_x_10")
      Appearance <- "DOx_Start_M_x_10"
   Button "Button_49" at 660,337 size 60x20; TextOff 'Выкл'; Authorization "Operate"
      on Click: ResetBit("DOx_Start_M_x_12")
      Appearance <- "DOx_Start_M_x_12"
   Button "Button_46" at 508,337 size 60x20; TextOff 'Выкл'; Authorization "Operate"
      on Click: ResetBit("DOx_Start_M_x_11")
      Appearance <- "DOx_Start_M_x_11"